   END_RUNG
   RUNG wire#w1
      Contact( #"TANK ACTIV 24" )
      Move(in := 3, out1 => #"GROUP of TANK 24")
   END_RUNG
   // the same network as SCL:
   IF #"SET GROUP 3" AND #"TANK ACTIV 1" THEN #"GROUP of TANK 1" := 3; END_IF;
   IF #"SET GROUP 3" AND #"TANK ACTIV 2" THEN #"GROUP of TANK 2" := 3; END_IF;
   IF #"SET GROUP 3" AND #"TANK ACTIV 3" THEN #"GROUP of TANK 3" := 3; END_IF;
   IF #"SET GROUP 3" AND #"TANK ACTIV 4" THEN #"GROUP of TANK 4" := 3; END_IF;
   IF #"SET GROUP 3" AND #"TANK ACTIV 5" THEN #"GROUP of TANK 5" := 3; END_IF;
   IF #"SET GROUP 3" AND #"TANK ACTIV 6" THEN #"GROUP of TANK 6" := 3; END_IF;
   IF #"SET GROUP 3" AND #"TANK ACTIV 7" THEN #"GROUP of TANK 7" := 3; END_IF;
   IF #"SET GROUP 3" AND #"TANK ACTIV 8" THEN #"GROUP of TANK 8" := 3; END_IF;
   IF #"SET GROUP 3" AND #"TANK ACTIV 9" THEN #"GROUP of TANK 9" := 3; END_IF;
   IF #"SET GROUP 3" AND #"TANK ACTIV 10" THEN #"GROUP of TANK 10" := 3; END_IF;
   IF #"SET GROUP 3" AND #"TANK ACTIV 11" THEN #"GROUP of TANK 11" := 3; END_IF;
   IF #"SET GROUP 3" AND #"TANK ACTIV 12" THEN #"GROUP of TANK 12" := 3; END_IF;
   IF #"SET GROUP 3" AND #"TANK ACTIV 13" THEN #"GROUP of TANK 13" := 3; END_IF;
   IF #"SET GROUP 3" AND #"TANK ACTIV 14" THEN #"GROUP of TANK 14" := 3; END_IF;
   IF #"SET GROUP 3" AND #"TANK ACTIV 15" THEN #"GROUP of TANK 15" := 3; END_IF;
   IF #"SET GROUP 3" AND #"TANK ACTIV 16" THEN #"GROUP of TANK 16" := 3; END_IF;
   IF #"SET GROUP 3" AND #"TANK ACTIV 17" THEN #"GROUP of TANK 17" := 3; END_IF;
   IF #"SET GROUP 3" AND #"TANK ACTIV 18" THEN #"GROUP of TANK 18" := 3; END_IF;
   IF #"SET GROUP 3" AND #"TANK ACTIV 19" THEN #"GROUP of TANK 19" := 3; END_IF;
   IF #"SET GROUP 3" AND #"TANK ACTIV 20" THEN #"GROUP of TANK 20" := 3; END_IF;
   IF #"SET GROUP 3" AND #"TANK ACTIV 21" THEN #"GROUP of TANK 21" := 3; END_IF;
   IF #"SET GROUP 3" AND #"TANK ACTIV 22" THEN #"GROUP of TANK 22" := 3; END_IF;
   IF #"SET GROUP 3" AND #"TANK ACTIV 23" THEN #"GROUP of TANK 23" := 3; END_IF;
   IF #"SET GROUP 3" AND #"TANK ACTIV 24" THEN #"GROUP of TANK 24" := 3; END_IF;
END_REGION

REGION Network 24: GROUP 4 of TANKS
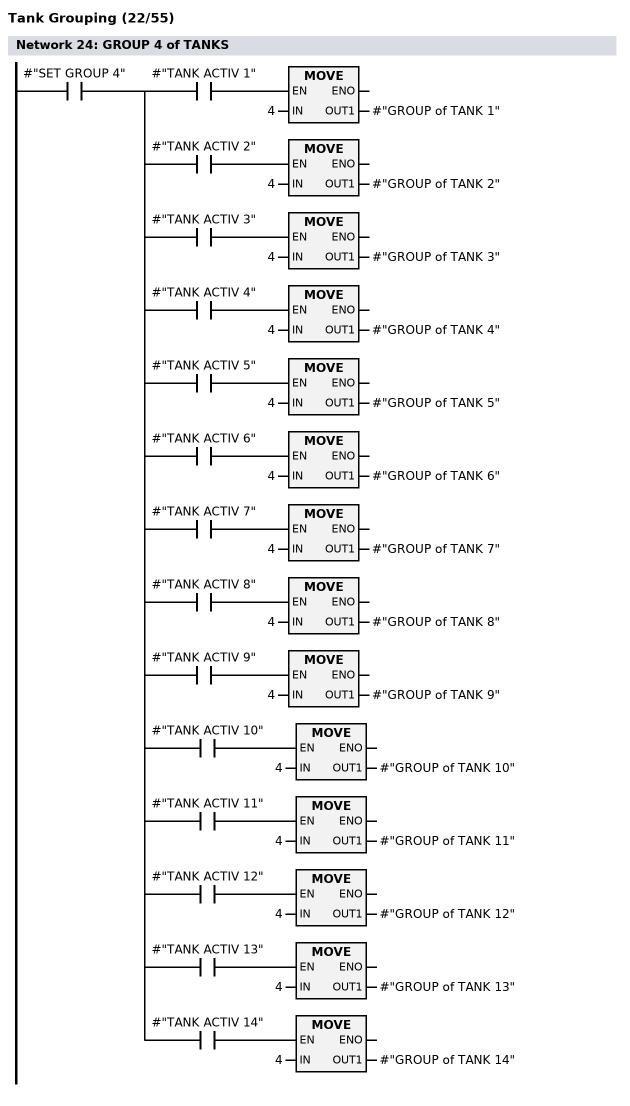
   RUNG wire#powerrail
      Contact( #"SET GROUP 4" )
      wire#w1
      Contact( #"TANK ACTIV 1" )
      Move(in := 4, out1 => #"GROUP of TANK 1")
   END_RUNG
   RUNG wire#w1
      Contact( #"TANK ACTIV 2" )
      Move(in := 4, out1 => #"GROUP of TANK 2")
   END_RUNG
   RUNG wire#w1
      Contact( #"TANK ACTIV 3" )
      Move(in := 4, out1 => #"GROUP of TANK 3")
   END_RUNG
   RUNG wire#w1
      Contact( #"TANK ACTIV 4" )
      Move(in := 4, out1 => #"GROUP of TANK 4")
   END_RUNG
   RUNG wire#w1
      Contact( #"TANK ACTIV 5" )
      Move(in := 4, out1 => #"GROUP of TANK 5")
   END_RUNG
   RUNG wire#w1
      Contact( #"TANK ACTIV 6" )
      Move(in := 4, out1 => #"GROUP of TANK 6")
   END_RUNG
   RUNG wire#w1
      Contact( #"TANK ACTIV 7" )
      Move(in := 4, out1 => #"GROUP of TANK 7")
   END_RUNG
   RUNG wire#w1
      Contact( #"TANK ACTIV 8" )
      Move(in := 4, out1 => #"GROUP of TANK 8")
   END_RUNG
   RUNG wire#w1
      Contact( #"TANK ACTIV 9" )
      Move(in := 4, out1 => #"GROUP of TANK 9")
   END_RUNG
   RUNG wire#w1
      Contact( #"TANK ACTIV 10" )
      Move(in := 4, out1 => #"GROUP of TANK 10")
   END_RUNG
   RUNG wire#w1
      Contact( #"TANK ACTIV 11" )
      Move(in := 4, out1 => #"GROUP of TANK 11")
   END_RUNG
   RUNG wire#w1
      Contact( #"TANK ACTIV 12" )
      Move(in := 4, out1 => #"GROUP of TANK 12")
   END_RUNG
   RUNG wire#w1
      Contact( #"TANK ACTIV 13" )
      Move(in := 4, out1 => #"GROUP of TANK 13")
   END_RUNG
   RUNG wire#w1
      Contact( #"TANK ACTIV 14" )
      Move(in := 4, out1 => #"GROUP of TANK 14")
   END_RUNG
   // the same network as SCL:
   IF #"SET GROUP 4" AND #"TANK ACTIV 1" THEN #"GROUP of TANK 1" := 4; END_IF;
   IF #"SET GROUP 4" AND #"TANK ACTIV 2" THEN #"GROUP of TANK 2" := 4; END_IF;
   IF #"SET GROUP 4" AND #"TANK ACTIV 3" THEN #"GROUP of TANK 3" := 4; END_IF;
   IF #"SET GROUP 4" AND #"TANK ACTIV 4" THEN #"GROUP of TANK 4" := 4; END_IF;
   IF #"SET GROUP 4" AND #"TANK ACTIV 5" THEN #"GROUP of TANK 5" := 4; END_IF;
   IF #"SET GROUP 4" AND #"TANK ACTIV 6" THEN #"GROUP of TANK 6" := 4; END_IF;
   IF #"SET GROUP 4" AND #"TANK ACTIV 7" THEN #"GROUP of TANK 7" := 4; END_IF;
   IF #"SET GROUP 4" AND #"TANK ACTIV 8" THEN #"GROUP of TANK 8" := 4; END_IF;
   IF #"SET GROUP 4" AND #"TANK ACTIV 9" THEN #"GROUP of TANK 9" := 4; END_IF;
   IF #"SET GROUP 4" AND #"TANK ACTIV 10" THEN #"GROUP of TANK 10" := 4; END_IF;
   IF #"SET GROUP 4" AND #"TANK ACTIV 11" THEN #"GROUP of TANK 11" := 4; END_IF;
   IF #"SET GROUP 4" AND #"TANK ACTIV 12" THEN #"GROUP of TANK 12" := 4; END_IF;
   IF #"SET GROUP 4" AND #"TANK ACTIV 13" THEN #"GROUP of TANK 13" := 4; END_IF;
   IF #"SET GROUP 4" AND #"TANK ACTIV 14" THEN #"GROUP of TANK 14" := 4; END_IF;
END_REGION

REGION Network 25: GROUP 5 of TANKS
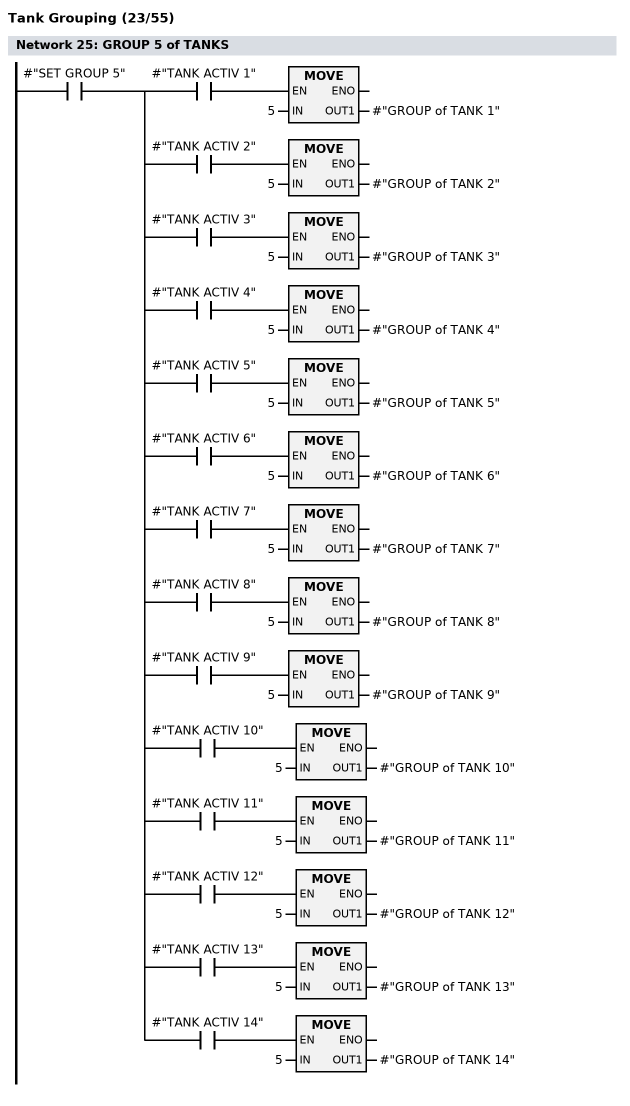
   RUNG wire#powerrail
      Contact( #"SET GROUP 5" )
      wire#w1
      Contact( #"TANK ACTIV 1" )
      Move(in := 5, out1 => #"GROUP of TANK 1")
   END_RUNG
   RUNG wire#w1
      Contact( #"TANK ACTIV 2" )
      Move(in := 5, out1 => #"GROUP of TANK 2")
   END_RUNG
   RUNG wire#w1
      Contact( #"TANK ACTIV 3" )
      Move(in := 5, out1 => #"GROUP of TANK 3")
   END_RUNG
   RUNG wire#w1
      Contact( #"TANK ACTIV 4" )
      Move(in := 5, out1 => #"GROUP of TANK 4")
   END_RUNG
   RUNG wire#w1
      Contact( #"TANK ACTIV 5" )
      Move(in := 5, out1 => #"GROUP of TANK 5")
   END_RUNG
   RUNG wire#w1
      Contact( #"TANK ACTIV 6" )
      Move(in := 5, out1 => #"GROUP of TANK 6")
   END_RUNG
   RUNG wire#w1
      Contact( #"TANK ACTIV 7" )
      Move(in := 5, out1 => #"GROUP of TANK 7")
   END_RUNG
   RUNG wire#w1
      Contact( #"TANK ACTIV 8" )
      Move(in := 5, out1 => #"GROUP of TANK 8")
   END_RUNG
   RUNG wire#w1
      Contact( #"TANK ACTIV 9" )
      Move(in := 5, out1 => #"GROUP of TANK 9")
   END_RUNG
   RUNG wire#w1
      Contact( #"TANK ACTIV 10" )
      Move(in := 5, out1 => #"GROUP of TANK 10")
   END_RUNG
   RUNG wire#w1
      Contact( #"TANK ACTIV 11" )
      Move(in := 5, out1 => #"GROUP of TANK 11")
   END_RUNG
   RUNG wire#w1
      Contact( #"TANK ACTIV 12" )
      Move(in := 5, out1 => #"GROUP of TANK 12")
   END_RUNG
   RUNG wire#w1
      Contact( #"TANK ACTIV 13" )
      Move(in := 5, out1 => #"GROUP of TANK 13")
   END_RUNG
   RUNG wire#w1
      Contact( #"TANK ACTIV 14" )
      Move(in := 5, out1 => #"GROUP of TANK 14")
   END_RUNG
   // the same network as SCL:
   IF #"SET GROUP 5" AND #"TANK ACTIV 1" THEN #"GROUP of TANK 1" := 5; END_IF;
   IF #"SET GROUP 5" AND #"TANK ACTIV 2" THEN #"GROUP of TANK 2" := 5; END_IF;
   IF #"SET GROUP 5" AND #"TANK ACTIV 3" THEN #"GROUP of TANK 3" := 5; END_IF;
   IF #"SET GROUP 5" AND #"TANK ACTIV 4" THEN #"GROUP of TANK 4" := 5; END_IF;
   IF #"SET GROUP 5" AND #"TANK ACTIV 5" THEN #"GROUP of TANK 5" := 5; END_IF;
   IF #"SET GROUP 5" AND #"TANK ACTIV 6" THEN #"GROUP of TANK 6" := 5; END_IF;
   IF #"SET GROUP 5" AND #"TANK ACTIV 7" THEN #"GROUP of TANK 7" := 5; END_IF;
   IF #"SET GROUP 5" AND #"TANK ACTIV 8" THEN #"GROUP of TANK 8" := 5; END_IF;
   IF #"SET GROUP 5" AND #"TANK ACTIV 9" THEN #"GROUP of TANK 9" := 5; END_IF;
   IF #"SET GROUP 5" AND #"TANK ACTIV 10" THEN #"GROUP of TANK 10" := 5; END_IF;
   IF #"SET GROUP 5" AND #"TANK ACTIV 11" THEN #"GROUP of TANK 11" := 5; END_IF;
   IF #"SET GROUP 5" AND #"TANK ACTIV 12" THEN #"GROUP of TANK 12" := 5; END_IF;
   IF #"SET GROUP 5" AND #"TANK ACTIV 13" THEN #"GROUP of TANK 13" := 5; END_IF;
   IF #"SET GROUP 5" AND #"TANK ACTIV 14" THEN #"GROUP of TANK 14" := 5; END_IF;
END_REGION

REGION Network 26: GROUP 6 of TANKS
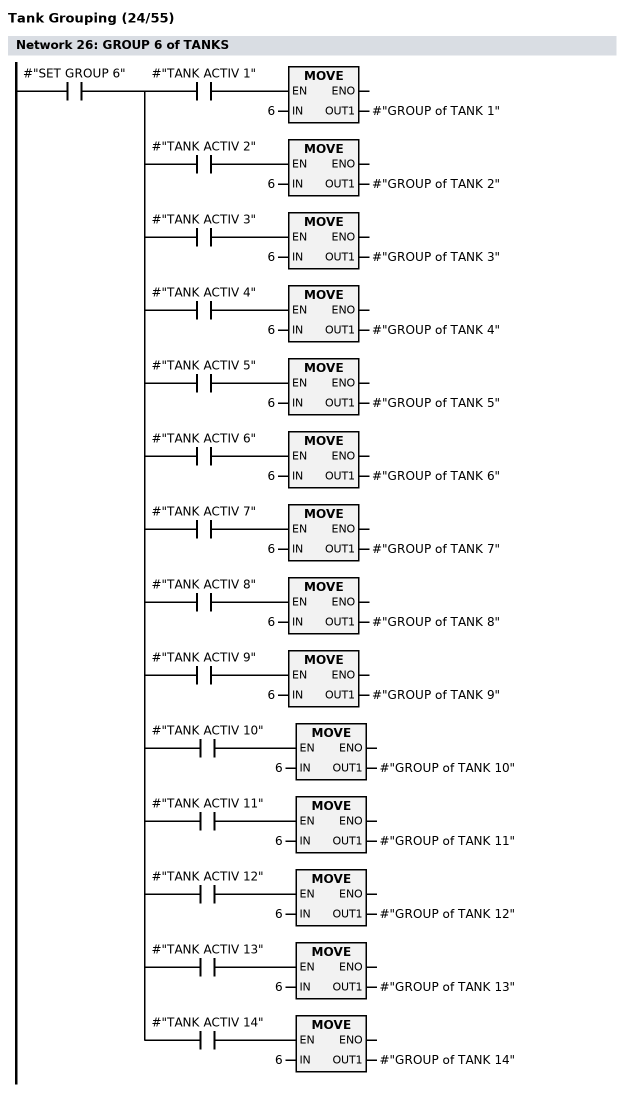
   RUNG wire#powerrail
      Contact( #"SET GROUP 6" )
      wire#w1
      Contact( #"TANK ACTIV 1" )
      Move(in := 6, out1 => #"GROUP of TANK 1")
   END_RUNG
   RUNG wire#w1
      Contact( #"TANK ACTIV 2" )
      Move(in := 6, out1 => #"GROUP of TANK 2")
   END_RUNG
   RUNG wire#w1
      Contact( #"TANK ACTIV 3" )
      Move(in := 6, out1 => #"GROUP of TANK 3")
   END_RUNG
   RUNG wire#w1
      Contact( #"TANK ACTIV 4" )
      Move(in := 6, out1 => #"GROUP of TANK 4")
   END_RUNG
   RUNG wire#w1
      Contact( #"TANK ACTIV 5" )
      Move(in := 6, out1 => #"GROUP of TANK 5")
   END_RUNG
   RUNG wire#w1
      Contact( #"TANK ACTIV 6" )
      Move(in := 6, out1 => #"GROUP of TANK 6")
   END_RUNG
   RUNG wire#w1
      Contact( #"TANK ACTIV 7" )
      Move(in := 6, out1 => #"GROUP of TANK 7")
   END_RUNG
   RUNG wire#w1
      Contact( #"TANK ACTIV 8" )
      Move(in := 6, out1 => #"GROUP of TANK 8")
   END_RUNG
   RUNG wire#w1
      Contact( #"TANK ACTIV 9" )
      Move(in := 6, out1 => #"GROUP of TANK 9")
   END_RUNG
   RUNG wire#w1
      Contact( #"TANK ACTIV 10" )
      Move(in := 6, out1 => #"GROUP of TANK 10")
   END_RUNG
   RUNG wire#w1
      Contact( #"TANK ACTIV 11" )
      Move(in := 6, out1 => #"GROUP of TANK 11")
   END_RUNG
   RUNG wire#w1
      Contact( #"TANK ACTIV 12" )
      Move(in := 6, out1 => #"GROUP of TANK 12")
   END_RUNG
   RUNG wire#w1
      Contact( #"TANK ACTIV 13" )
      Move(in := 6, out1 => #"GROUP of TANK 13")
   END_RUNG
   RUNG wire#w1
      Contact( #"TANK ACTIV 14" )
      Move(in := 6, out1 => #"GROUP of TANK 14")
   END_RUNG
   // the same network as SCL:
   IF #"SET GROUP 6" AND #"TANK ACTIV 1" THEN #"GROUP of TANK 1" := 6; END_IF;
   IF #"SET GROUP 6" AND #"TANK ACTIV 2" THEN #"GROUP of TANK 2" := 6; END_IF;
   IF #"SET GROUP 6" AND #"TANK ACTIV 3" THEN #"GROUP of TANK 3" := 6; END_IF;
   IF #"SET GROUP 6" AND #"TANK ACTIV 4" THEN #"GROUP of TANK 4" := 6; END_IF;
   IF #"SET GROUP 6" AND #"TANK ACTIV 5" THEN #"GROUP of TANK 5" := 6; END_IF;
   IF #"SET GROUP 6" AND #"TANK ACTIV 6" THEN #"GROUP of TANK 6" := 6; END_IF;
   IF #"SET GROUP 6" AND #"TANK ACTIV 7" THEN #"GROUP of TANK 7" := 6; END_IF;
   IF #"SET GROUP 6" AND #"TANK ACTIV 8" THEN #"GROUP of TANK 8" := 6; END_IF;
   IF #"SET GROUP 6" AND #"TANK ACTIV 9" THEN #"GROUP of TANK 9" := 6; END_IF;
   IF #"SET GROUP 6" AND #"TANK ACTIV 10" THEN #"GROUP of TANK 10" := 6; END_IF;
   IF #"SET GROUP 6" AND #"TANK ACTIV 11" THEN #"GROUP of TANK 11" := 6; END_IF;
   IF #"SET GROUP 6" AND #"TANK ACTIV 12" THEN #"GROUP of TANK 12" := 6; END_IF;
   IF #"SET GROUP 6" AND #"TANK ACTIV 13" THEN #"GROUP of TANK 13" := 6; END_IF;
   IF #"SET GROUP 6" AND #"TANK ACTIV 14" THEN #"GROUP of TANK 14" := 6; END_IF;
END_REGION

REGION Network 27: GROUP 7 of TANKS
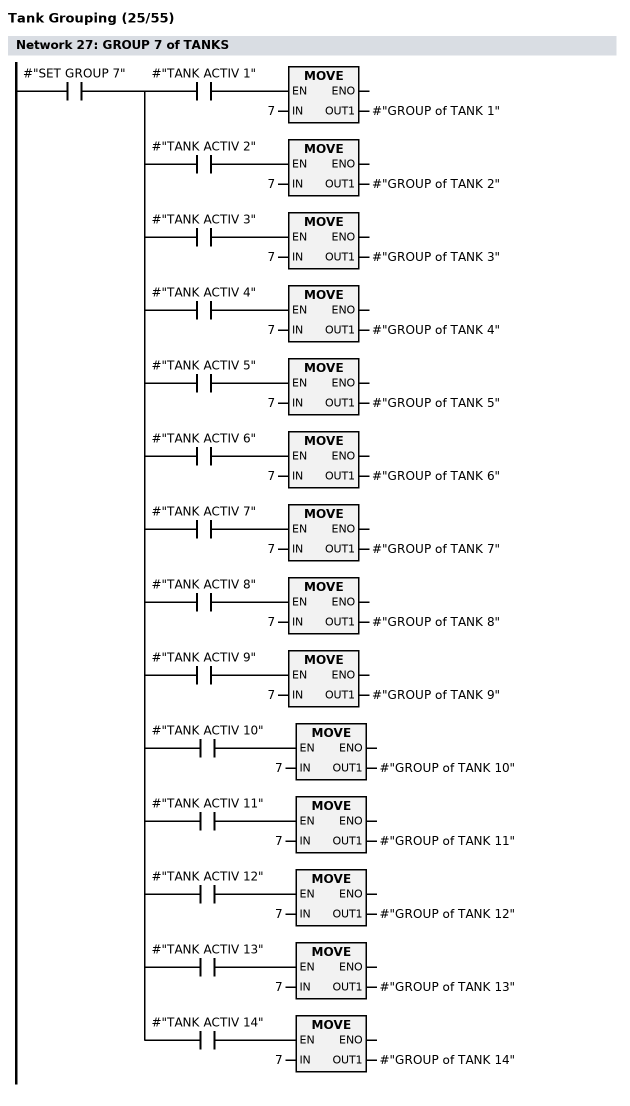
   RUNG wire#powerrail
      Contact( #"SET GROUP 7" )
      wire#w1
      Contact( #"TANK ACTIV 1" )
      Move(in := 7, out1 => #"GROUP of TANK 1")
   END_RUNG
   RUNG wire#w1
      Contact( #"TANK ACTIV 2" )
      Move(in := 7, out1 => #"GROUP of TANK 2")
   END_RUNG
   RUNG wire#w1
      Contact( #"TANK ACTIV 3" )
      Move(in := 7, out1 => #"GROUP of TANK 3")
   END_RUNG
   RUNG wire#w1
      Contact( #"TANK ACTIV 4" )
      Move(in := 7, out1 => #"GROUP of TANK 4")
   END_RUNG
   RUNG wire#w1
      Contact( #"TANK ACTIV 5" )
      Move(in := 7, out1 => #"GROUP of TANK 5")
   END_RUNG
   RUNG wire#w1
      Contact( #"TANK ACTIV 6" )
      Move(in := 7, out1 => #"GROUP of TANK 6")
   END_RUNG
   RUNG wire#w1
      Contact( #"TANK ACTIV 7" )
      Move(in := 7, out1 => #"GROUP of TANK 7")
   END_RUNG
   RUNG wire#w1
      Contact( #"TANK ACTIV 8" )
      Move(in := 7, out1 => #"GROUP of TANK 8")
   END_RUNG
   RUNG wire#w1
      Contact( #"TANK ACTIV 9" )
      Move(in := 7, out1 => #"GROUP of TANK 9")
   END_RUNG
   RUNG wire#w1
      Contact( #"TANK ACTIV 10" )
      Move(in := 7, out1 => #"GROUP of TANK 10")
   END_RUNG
   RUNG wire#w1
      Contact( #"TANK ACTIV 11" )
      Move(in := 7, out1 => #"GROUP of TANK 11")
   END_RUNG
   RUNG wire#w1
      Contact( #"TANK ACTIV 12" )
      Move(in := 7, out1 => #"GROUP of TANK 12")
   END_RUNG
   RUNG wire#w1
      Contact( #"TANK ACTIV 13" )
      Move(in := 7, out1 => #"GROUP of TANK 13")
   END_RUNG
   RUNG wire#w1
      Contact( #"TANK ACTIV 14" )
      Move(in := 7, out1 => #"GROUP of TANK 14")
   END_RUNG
   // the same network as SCL:
   IF #"SET GROUP 7" AND #"TANK ACTIV 1" THEN #"GROUP of TANK 1" := 7; END_IF;
   IF #"SET GROUP 7" AND #"TANK ACTIV 2" THEN #"GROUP of TANK 2" := 7; END_IF;
   IF #"SET GROUP 7" AND #"TANK ACTIV 3" THEN #"GROUP of TANK 3" := 7; END_IF;
   IF #"SET GROUP 7" AND #"TANK ACTIV 4" THEN #"GROUP of TANK 4" := 7; END_IF;
   IF #"SET GROUP 7" AND #"TANK ACTIV 5" THEN #"GROUP of TANK 5" := 7; END_IF;
   IF #"SET GROUP 7" AND #"TANK ACTIV 6" THEN #"GROUP of TANK 6" := 7; END_IF;
   IF #"SET GROUP 7" AND #"TANK ACTIV 7" THEN #"GROUP of TANK 7" := 7; END_IF;
   IF #"SET GROUP 7" AND #"TANK ACTIV 8" THEN #"GROUP of TANK 8" := 7; END_IF;
   IF #"SET GROUP 7" AND #"TANK ACTIV 9" THEN #"GROUP of TANK 9" := 7; END_IF;
   IF #"SET GROUP 7" AND #"TANK ACTIV 10" THEN #"GROUP of TANK 10" := 7; END_IF;
   IF #"SET GROUP 7" AND #"TANK ACTIV 11" THEN #"GROUP of TANK 11" := 7; END_IF;
   IF #"SET GROUP 7" AND #"TANK ACTIV 12" THEN #"GROUP of TANK 12" := 7; END_IF;
   IF #"SET GROUP 7" AND #"TANK ACTIV 13" THEN #"GROUP of TANK 13" := 7; END_IF;
   IF #"SET GROUP 7" AND #"TANK ACTIV 14" THEN #"GROUP of TANK 14" := 7; END_IF;
END_REGION

REGION Network 28: GROUP 8 of TANKS
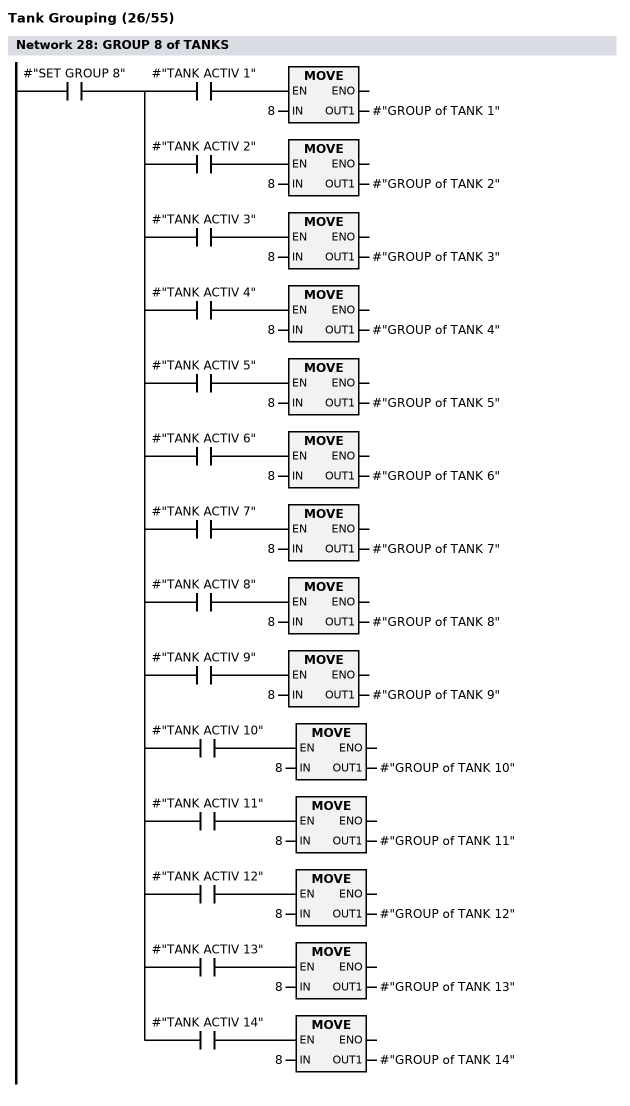
   RUNG wire#powerrail
      Contact( #"SET GROUP 8" )
      wire#w1
      Contact( #"TANK ACTIV 1" )
      Move(in := 8, out1 => #"GROUP of TANK 1")
   END_RUNG
   RUNG wire#w1
      Contact( #"TANK ACTIV 2" )
      Move(in := 8, out1 => #"GROUP of TANK 2")
   END_RUNG
   RUNG wire#w1
      Contact( #"TANK ACTIV 3" )
      Move(in := 8, out1 => #"GROUP of TANK 3")
   END_RUNG
   RUNG wire#w1
      Contact( #"TANK ACTIV 4" )
      Move(in := 8, out1 => #"GROUP of TANK 4")
   END_RUNG
   RUNG wire#w1
      Contact( #"TANK ACTIV 5" )
      Move(in := 8, out1 => #"GROUP of TANK 5")
   END_RUNG
   RUNG wire#w1
      Contact( #"TANK ACTIV 6" )
      Move(in := 8, out1 => #"GROUP of TANK 6")
   END_RUNG
   RUNG wire#w1
      Contact( #"TANK ACTIV 7" )
      Move(in := 8, out1 => #"GROUP of TANK 7")
   END_RUNG
   RUNG wire#w1
      Contact( #"TANK ACTIV 8" )
      Move(in := 8, out1 => #"GROUP of TANK 8")
   END_RUNG
   RUNG wire#w1
      Contact( #"TANK ACTIV 9" )
      Move(in := 8, out1 => #"GROUP of TANK 9")
   END_RUNG
   RUNG wire#w1
      Contact( #"TANK ACTIV 10" )
      Move(in := 8, out1 => #"GROUP of TANK 10")
   END_RUNG
   RUNG wire#w1
      Contact( #"TANK ACTIV 11" )
      Move(in := 8, out1 => #"GROUP of TANK 11")
   END_RUNG
   RUNG wire#w1
      Contact( #"TANK ACTIV 12" )
      Move(in := 8, out1 => #"GROUP of TANK 12")
   END_RUNG
   RUNG wire#w1
      Contact( #"TANK ACTIV 13" )
      Move(in := 8, out1 => #"GROUP of TANK 13")
   END_RUNG
   RUNG wire#w1
      Contact( #"TANK ACTIV 14" )
      Move(in := 8, out1 => #"GROUP of TANK 14")
   END_RUNG
   // the same network as SCL:
   IF #"SET GROUP 8" AND #"TANK ACTIV 1" THEN #"GROUP of TANK 1" := 8; END_IF;
   IF #"SET GROUP 8" AND #"TANK ACTIV 2" THEN #"GROUP of TANK 2" := 8; END_IF;
   IF #"SET GROUP 8" AND #"TANK ACTIV 3" THEN #"GROUP of TANK 3" := 8; END_IF;
   IF #"SET GROUP 8" AND #"TANK ACTIV 4" THEN #"GROUP of TANK 4" := 8; END_IF;
   IF #"SET GROUP 8" AND #"TANK ACTIV 5" THEN #"GROUP of TANK 5" := 8; END_IF;
   IF #"SET GROUP 8" AND #"TANK ACTIV 6" THEN #"GROUP of TANK 6" := 8; END_IF;
   IF #"SET GROUP 8" AND #"TANK ACTIV 7" THEN #"GROUP of TANK 7" := 8; END_IF;
   IF #"SET GROUP 8" AND #"TANK ACTIV 8" THEN #"GROUP of TANK 8" := 8; END_IF;
   IF #"SET GROUP 8" AND #"TANK ACTIV 9" THEN #"GROUP of TANK 9" := 8; END_IF;
   IF #"SET GROUP 8" AND #"TANK ACTIV 10" THEN #"GROUP of TANK 10" := 8; END_IF;
   IF #"SET GROUP 8" AND #"TANK ACTIV 11" THEN #"GROUP of TANK 11" := 8; END_IF;
   IF #"SET GROUP 8" AND #"TANK ACTIV 12" THEN #"GROUP of TANK 12" := 8; END_IF;
   IF #"SET GROUP 8" AND #"TANK ACTIV 13" THEN #"GROUP of TANK 13" := 8; END_IF;
   IF #"SET GROUP 8" AND #"TANK ACTIV 14" THEN #"GROUP of TANK 14" := 8; END_IF;
END_REGION

REGION Network 29: GROUP 9 of TANKS
